// TIA Portal project "Factory_Project_V17" (V17)
// Vorlageprojekt für das Buch mit Zielsystem S7-1200

(* hardware
DEVICE "S7-1200-Station_1"  S7-1200 Station
   slot 0: "Baugruppenträger_0"  Rack  V1.0
   slot 1: "PLC_1"  CPU 1211C DC/DC/DC  6ES7 211-1AE40-0XB0  V4.1
DEVICE "HMI_1"  KTP700 Basic PN
   slot 0: "HMI_1"  KTP700 Basic PN  6AV2 123-2GB03-0AX0  17.0.0.0
   slot 1: "HMI_RT_1"  KTP700 Basic PN  6AV2 123-2GB03-0AX0  17.0.0.0
   slot 5: "HMI_1.IE_CP_1"  PROFINET Interface  17.0.0.0
      slot 1: "PROFINET Interface_1"  PROFINET Interface
         slot 1: "Port_1"  Port
*)

// ===== PLC "PLC_1"  CPU 1211C DC/DC/DC =====

VAR_GLOBAL   // PLC tag table "Standard-Variablentabelle"
   "Tag_4" AT %M0.0 : Bool;
   "Tag_5" AT %M0.1 : Bool;
   "Tag_1" AT %M0.3 : Bool;
   "Tag_2" AT %M0.4 : Bool;
   "Tag_3" AT %M100.0 : Bool;
   "Tag_6" AT %M100.1 : Bool;
   "Tag_7" AT %M100.2 : Bool;
   "Tag_8" AT %M100.3 : Bool;
   "Tag_9" AT %M100.4 : Bool;
   "Tag_10" AT %M100.5 : Bool;
   "Tag_11" AT %M100.6 : Bool;
   "Tag_12" AT %M100.7 : Bool;
END_VAR

VAR_GLOBAL   // PLC tag table "Inputs_Tags"
   "start" AT %I0.0 : Bool;
   "stop" AT %I0.1 : Bool;
   "reset" AT %I0.2 : Bool;
   "emergency" AT %I0.3 : Bool;
   "Z1_Presence_sensor" AT %I0.4 : Bool;
   "at_scale_sensor" AT %I0.5 : Bool;
   "Z1_vision_sensor" AT %I0.6 : Bool;
   "machine A entry sensor" AT %I0.7 : Bool;
   "machine B entry sensor" AT %I1.0 : Bool;
   "machine A exit sensor" AT %I1.1 : Bool;
   "machine B exit sensor" AT %I1.2 : Bool;
   "machine A has error" AT %I1.3 : Bool;
   "machine A is busy" AT %I1.4 : Bool;
   "machine A opened" AT %I1.5 : Bool;
   "machine B has error" AT %I1.6 : Bool;
   "machine B is busy" AT %I1.7 : Bool;
   "machine B opened" AT %I2.0 : Bool;
   "up elevator A right limit" AT %I2.1 : Bool;
   "up elevator A left limit" AT %I2.2 : Bool;
   "down elevator A right limit" AT %I2.3 : Bool;
   "down elevator A left limit" AT %I2.4 : Bool;
   "up elevator B right limit" AT %I2.5 : Bool;
   "up elevator B left limit" AT %I2.6 : Bool;
   "down elevator B right limit" AT %I2.7 : Bool;
   "down elevator B left limit" AT %I3.0 : Bool;
   "product A at assemply" AT %I3.3 : Bool;
   "product B at assemply" AT %I3.4 : Bool;
   "product left assemply" AT %I3.5 : Bool;
   "positioner A limit" AT %I3.6 : Bool;
   "positioner A clamped" AT %I3.7 : Bool;
   "positioner B limit" AT %I4.0 : Bool;
   "Positioner B clamped" AT %I4.1 : Bool;
   "assempler moving x" AT %I4.2 : Bool;
   "assempler  moving z" AT %I4.3 : Bool;
   "assempler rotating" AT %I4.4 : Bool;
   "assempler item detected" AT %I4.5 : Bool;
   "assempler gripper rotating" AT %I4.6 : Bool;
   "palletizer elevator back limit" AT %I4.7 : Bool;
   "palletizer elevator front limit" AT %I5.0 : Bool;
   "palletizer clamped" AT %I5.1 : Bool;
   "palletizer elevator moving" AT %I5.2 : Bool;
   "palletizer plate limit" AT %I5.3 : Bool;
   "palletizer pusher limit" AT %I5.4 : Bool;
   "stacker crane moving x" AT %I5.5 : Bool;
   "stacker crane moving z" AT %I5.6 : Bool;
   "stacker crane left limit" AT %I5.7 : Bool;
   "stacker crane right limit" AT %I6.0 : Bool;
   "stacker crane middle limit" AT %I6.1 : Bool;
   "scale value" AT %ID32 : Real;
   "UP ELEVATOR A POSITION" AT %ID36 : Real;
   "DOWN ELEVATOR A POSITION" AT %ID40 : Real;
   "assempler position x" AT %ID44 : Real;
   "assempler position z" AT %ID48 : Real;
   "bridge A1 sensor" AT %I6.2 : Bool;
   "bridge A2 sensor" AT %I6.3 : Bool;
   "bridge B1 sensor" AT %I6.4 : Bool;
   "bridge B2 sensor" AT %I6.5 : Bool;
   "UP ELEVATOR B POSITION" AT %ID52 : Real;
   "DOWN ELEVATOR B POSITION" AT %ID56 : Real;
   "PALLETIZER ENTRY" AT %I6.6 : Bool;
   "LOADING CONV ENTRY SENSOR" AT %I6.7 : Bool;
   "LOADING CONV EXIT SENSOR" AT %I7.0 : Bool;
END_VAR

VAR_GLOBAL   // PLC tag table "Outputs_tags"
   "start light" AT %Q0.0 : Bool;
   "stop light" AT %Q0.1 : Bool;
   "reset light" AT %Q0.2 : Bool;
   "error light 1" AT %Q0.3 : Bool;
   "error light 2" AT %Q0.4 : Bool;
   "warning light 1" AT %Q0.5 : Bool;
   "warning light 2" AT %Q0.6 : Bool;
   "feed conv" AT %Q0.7 : Bool;
   "feed emittor" AT %Q1.0 : Bool;
   "scale conv" AT %Q1.1 : Bool;
   "sorter wheels" AT %Q1.2 : Bool;
   "sorter right" AT %Q1.3 : Bool;
   "sorter left" AT %Q1.4 : Bool;
   "Z1L1" AT %Q1.5 : Bool;
   "Z1L2" AT %Q1.6 : Bool;
   "Z1L3" AT %Q1.7 : Bool;
   "Z1L4" AT %Q2.0 : Bool;
   "Z1L5" AT %Q2.1 : Bool;
   "Z1L6" AT %Q2.2 : Bool;
   "Z1L7" AT %Q2.3 : Bool;
   "Z1L8" AT %Q2.4 : Bool;
   "Z1R1" AT %Q2.5 : Bool;
   "Z1R2" AT %Q2.6 : Bool;
   "Z1R3" AT %Q2.7 : Bool;
   "Z1R4" AT %Q3.0 : Bool;
   "Z1R5" AT %Q3.1 : Bool;
   "Z1R6" AT %Q3.2 : Bool;
   "Z3A1" AT %Q3.3 : Bool;
   "Z3A2" AT %Q3.4 : Bool;
   "Z3A3" AT %Q3.5 : Bool;
   "Z3A4" AT %Q3.6 : Bool;
   "Z3A5" AT %Q3.7 : Bool;
   "Z3A6" AT %Q4.0 : Bool;
   "Z3B1" AT %Q4.1 : Bool;
   "Z3B2" AT %Q4.2 : Bool;
   "Z3B3" AT %Q4.3 : Bool;
   "Z3B4" AT %Q4.4 : Bool;
   "Z3B5" AT %Q4.5 : Bool;
   "Z3B6" AT %Q4.6 : Bool;
   "Z3B7" AT %Q4.7 : Bool;
   "Z4_1" AT %Q5.2 : Bool;
   "Z4_2" AT %Q5.3 : Bool;
   "Z4_3" AT %Q5.4 : Bool;
   "Z4_4" AT %Q5.5 : Bool;
   "Z4 entry roller" AT %Q5.7 : Bool;
   "Z4 exit roller" AT %Q6.0 : Bool;
   "loading entry conv" AT %Q6.1 : Bool;
   "loading exit conv" AT %Q6.2 : Bool;
   "exit conv 1" AT %Q6.3 : Bool;
   "exit conv 2" AT %Q6.4 : Bool;
   "exit conv 3" AT %Q6.5 : Bool;
   "machine A start" AT %Q6.6 : Bool;
   "machine A stop" AT %Q6.7 : Bool;
   "machine A reset" AT %Q7.0 : Bool;
   "machine A lids" AT %Q7.1 : Bool;
   "machine B start" AT %Q7.2 : Bool;
   "Z4_5" AT %Q5.6 : Bool;
   "machine B stop" AT %Q7.3 : Bool;
   "machine B reset" AT %Q7.4 : Bool;
   "machine B lids" AT %Q7.5 : Bool;
   "up elevator A +" AT %Q7.6 : Bool;
   "up elevator A -" AT %Q7.7 : Bool;
   "up elevator A stop blade" AT %Q8.0 : Bool;
   "up elevator B +" AT %Q8.1 : Bool;
   "up elevator B -" AT %Q8.2 : Bool;
   "up elevator B stop blade" AT %Q8.3 : Bool;
   "down elevator A +" AT %Q8.4 : Bool;
   "down elevator A -" AT %Q8.5 : Bool;
   "down elevator A stop blade" AT %Q8.6 : Bool;
   "down elevator B+" AT %Q8.7 : Bool;
   "down elevator B -" AT %Q9.0 : Bool;
   "down elevator B stop blade" AT %Q9.1 : Bool;
   "positioner A raise" AT %Q9.2 : Bool;
   "positioner A clamp" AT %Q9.3 : Bool;
   "positioner B raise" AT %Q9.4 : Bool;
   "positioner B clamp" AT %Q9.5 : Bool;
   "assempler grap" AT %Q9.6 : Bool;
   "assempler rotate cw" AT %Q9.7 : Bool;
   "assempler rotate ccw" AT %Q10.1 : Bool;
   "assempler gripper ccw" AT %Q10.2 : Bool;
   "palletizer turn" AT %Q10.3 : Bool;
   "palletizer push" AT %Q10.4 : Bool;
   "palletizer clamp" AT %Q10.5 : Bool;
   "palletizer open plate" AT %Q10.6 : Bool;
   "palletizer belt +" AT %Q10.7 : Bool;
   "palletizer belt -" AT %Q11.0 : Bool;
   "palletizer chain +" AT %Q11.1 : Bool;
   "palletizer chain -" AT %Q11.2 : Bool;
   "palletizer elevator +" AT %Q11.3 : Bool;
   "palletizer elevator -" AT %Q11.4 : Bool;
   "palletizer elevator move to limit" AT %Q11.5 : Bool;
   "stacker crane lift" AT %Q11.6 : Bool;
   "stacker crane left" AT %Q11.7 : Bool;
   "stacker crane right" AT %Q12.0 : Bool;
   "state" AT %QD32 : DInt;
   "up elevator A set point" AT %QD36 : Real;
   "up elevator B set point" AT %QD40 : Real;
   "down elevator A set point" AT %QD44 : Real;
   "down elevator B set point" AT %QD48 : Real;
   "assempler x set point" AT %QD52 : Real;
   "assempler z set point" AT %QD56 : Real;
   "stacker crane target position" AT %QD60 : DInt;
   "bridge A1 stop blade" AT %Q12.1 : Bool;
   "bridge A2 stop blade" AT %Q12.2 : Bool;
   "bridge B1 stop blade" AT %Q12.3 : Bool;
   "bridge B2 stop blade" AT %Q12.4 : Bool;
   "Z3-A1 bridge conv" AT %Q12.5 : Bool;
   "Z3-A2 bridge conv" AT %Q12.6 : Bool;
   "Z3-A3 bridge conv" AT %Q12.7 : Bool;
   "Z3-B1 bridge conv" AT %Q13.0 : Bool;
   "Z3-B2 bridge conv" AT %Q13.1 : Bool;
   "Z3-B3 bridge conv" AT %Q13.2 : Bool;
   "PALLETIZER EMITTER" AT %Q10.0 : Bool;
END_VAR

VAR_GLOBAL   // PLC tag table "alarm_tags"
   "Alarm_trigger" AT %MW100 : Word;
END_VAR

TYPE "RackSlot"
   STRUCT
      occupied : Bool;
      side : Int;
      space : Int;
   END_STRUCT;
END_TYPE

DATA_BLOCK "DB_RackMemory"   // DB8
{ S7_Optimized_Access := 'TRUE' }
VERSION : 0.1
   VAR
      Rack : Array[1..108] of "RackSlot";
      SpacesOccupied : Int;
      "FREE SPACES" : Int;
      "QUANTITY TO RETRIEVE" : Int;
      "REQUIRED QUANTITY" : Int;
      RETRIEVE : Bool;
      In_Production : Int;
      "TOTAL ORDERS" : Int;
      "TOTAL DLIEVERED" : Int;
      ReckMemoryReset : Bool;
      InProductionReset : Bool;
   END_VAR
BEGIN
END_DATA_BLOCK

DATA_BLOCK "DB_HMI"   // DB10
{ S7_Optimized_Access := 'TRUE' }
VERSION : 0.1
   VAR
      "Z1 STATUS" : Int;
      "Z2 STATUS" : Int;
      "Z3 BUFFER A STATUS" : Int;
      "Z3 BUFFER B STATUS" : Int;
      "Z3 ASSEMPLER STATUS" : Int;
      "Z4 UPPER STATUS" : Int;
      "Z4 LOWER STATUS" : Int;
      "Z5 STATUS" : Int;
      "FACTORY STATUS" : Int;
      "ASSEMPLER X" : Real;
      "ASSEMPLER Z" : Real;
      "ASSEMPLER GRAB" : Bool;
      "ASSEMPLER ROT CW" : Bool;
      "ASSEMPLER ROT CCW" : Bool;
      "CRANE TARGET" : Int;
      "CRANE SIDE" : Int;
      "CRANE LEFT" : Bool;
      "CRANE LIFT" : Bool;
      "CRANE RIGHT" : Bool;
      "CREATE ORDER" : Bool;
      "CANCEL ORDER" : Bool;
      "MAINTENANCE MODE" : Bool;
      ACK : Bool;
   END_VAR
BEGIN
END_DATA_BLOCK

DATA_BLOCK "FACTORY STATUS MANAGMENT_DB"   // DB11
{ S7_Optimized_Access := 'TRUE' }
VERSION : 0.1
// stored: InstanceOfName FACTORY STATUS MANAGMENT
"FACTORY STATUS MANAGMENT"
BEGIN
END_DATA_BLOCK

// folder: System blocks/Program resources

DATA_BLOCK "z1_timer_ton"   // DB3
{ S7_Optimized_Access := 'TRUE' }
AUTHOR : Simatic
FAMILY : IEC
NAME : IEC_TMR
VERSION : 1.0
// stored: InstanceOfName IEC_TIMER
"IEC_TIMER"
BEGIN
END_DATA_BLOCK

// folder: ZONE-5-BLOCKS

DATA_BLOCK "ZONE-5-FB_DB"   // DB9
{ S7_Optimized_Access := 'TRUE' }
VERSION : 0.1
// stored: InstanceOfName ZONE-5-FB
"ZONE-5-FB"
BEGIN
END_DATA_BLOCK

// folder: ZONE_1_BLOCKS

DATA_BLOCK "Zone_1_FB_DB"   // DB2
{ S7_Optimized_Access := 'TRUE' }
VERSION : 0.1
// stored: InstanceOfName Zone_1_FB
"Zone_1_FB"
BEGIN
END_DATA_BLOCK

// folder: ZONE_4_BLOCKS

DATA_BLOCK "ZONE 4 FB_DB"   // DB7
{ S7_Optimized_Access := 'TRUE' }
VERSION : 0.1
// stored: InstanceOfName ZONE 4 FB
"ZONE 4 FB"
BEGIN
END_DATA_BLOCK

// folder: Zone _2_Blocks

DATA_BLOCK "Zone_2_FB_DB"   // DB4
{ S7_Optimized_Access := 'TRUE' }
VERSION : 0.1
// stored: InstanceOfName Zone_2_FB
"Zone_2_FB"
BEGIN
END_DATA_BLOCK

// folder: Zone_3_blocks

DATA_BLOCK "Zone_3_FB_DB"   // DB5
{ S7_Optimized_Access := 'TRUE' }
VERSION : 0.1
// stored: InstanceOfName Zone_3_FB
"Zone_3_FB"
BEGIN
END_DATA_BLOCK

// folder: Zone_3_blocks/BUFFER SUB BLOCKS

DATA_BLOCK "ZONE-3 BUFFER_A_DB"   // DB6
{ S7_Optimized_Access := 'TRUE' }
VERSION : 0.1
// stored: InstanceOfName ZONE-3 BUFFER
"ZONE-3 BUFFER"
BEGIN
END_DATA_BLOCK

// folder: (top level)

FUNCTION_BLOCK "FACTORY STATUS MANAGMENT"   // FB22, SCL
{ S7_Optimized_Access := 'TRUE' }
VERSION : 0.1
   VAR_INPUT
      START : Bool;
      STOP : Bool;
      RESET : Bool;
      "Z1 STATUS" : Int;
      "Z2 STATUS" : Int;
      "Z3 BUFFER A STATUS" : Int;
      "Z3 BUFFER B STATUS" : Int;
      "Z3 ASSEMPLER STATUS" : Int;
      "Z4 STATUS UPPER" : Int;
      "Z4 LOWER STATUS" : Int;
      "Z5 STATUS" : Int;
   END_VAR
   VAR_OUTPUT
      "FACTORY STATUS" : Int;
   END_VAR
BEGIN
   IF #"Z1 STATUS" = 90
       OR #"Z2 STATUS" = 90
       OR #"Z3 BUFFER A STATUS" = 90
       OR #"Z3 BUFFER B STATUS" = 90
       OR #"Z3 ASSEMPLER STATUS" = 90
       OR #"Z4 STATUS UPPER" = 90
       OR #"Z4 LOWER STATUS" = 90
       OR #"Z5 STATUS" = 90
   THEN
       #"FACTORY STATUS" := 90;
   END_IF;

   IF #"FACTORY STATUS" = 90 THEN
       IF #RESET THEN
           #"FACTORY STATUS" := 0;
       END_IF;
   END_IF;

   IF #START AND  #"FACTORY STATUS" <> 90 THEN
       #"FACTORY STATUS" := 10;
   END_IF;

   IF #STOP AND #"FACTORY STATUS" <> 90 THEN
       #"FACTORY STATUS" := 0;
   END_IF;
END_FUNCTION_BLOCK

FUNCTION "MHJ-PLC-Lab-Function-S71200" : Void   // FC9000, SCL
{ S7_Optimized_Access := 'TRUE' }
VERSION : 0.1
   VAR_TEMP
      rdTimeReturn : Int;
      outputTime : DTL;
      SyncVal : Byte;
      forVal : Int;
      forVal_2 : Int;
      Value : Byte;
   END_VAR
   VAR CONSTANT
      CompVal : Byte := 16#34;
      Value_01 : Byte := 16#11;
      Value_01_DW : DWord := 16#A165_D992;
      Value_02_DW : DWord := 16#58BE_4401;
   END_VAR
BEGIN

   #Value:=PEEK(area := 16#82,
        dbNumber := 0,
        byteOffset := 511);
   #Value := #Value + 1;

   POKE(area := 16#82,
        dbNumber := 0,
        byteOffset := 511,
        value := #Value);

   POKE(area:=16#81,
        dbNumber:=0,
        byteOffset:=1016,
        value:=#Value_01_DW);
   POKE(area := 16#81,
        dbNumber := 0,
        byteOffset := 1020,
        value := #Value_02_DW);

   POKE(area := 16#81,
        dbNumber := 0,
        byteOffset := 511,
        value := B#16#00);

   FOR #forVal := 0 TO 120 DO
       FOR #forVal_2:=0 TO 10 DO
           #rdTimeReturn:=RD_SYS_T(#outputTime);
           #rdTimeReturn := WR_SYS_T(#outputTime);
           #rdTimeReturn := RD_SYS_T(#outputTime);
           #rdTimeReturn := WR_SYS_T(#outputTime);
       END_FOR;
       #SyncVal:= PEEK(area := 16#81,
                      dbNumber := 0,
                      byteOffset := 511);
       IF #SyncVal = #CompVal THEN
          GOTO M_1;
       END_IF;
   END_FOR;
   RETURN;

   M_1:
   POKE(area := 16#81,
        dbNumber := 0,
        byteOffset := 511,
        value := B#16#0);
END_FUNCTION

ORGANIZATION_BLOCK "Main"   // OB1, LAD, ProgramCycle
TITLE = "Main Program Sweep (Cycle)"
{ S7_Optimized_Access := 'TRUE' }
VERSION : 0.1
   VAR_INPUT
      Initial_Call : Bool;   // Initial call of this OB
      Remanence : Bool;   // =True, if remanent data are available
   END_VAR
BEGIN

REGION Network 1: Konnektierungsbaustein für PLC-Lab
   // Im Netzwerk 1 wird der Konnektierungsbaustein für PLC-Lab aufgerufen.
   // Dieser Aufruf darf nicht entfernt werden!
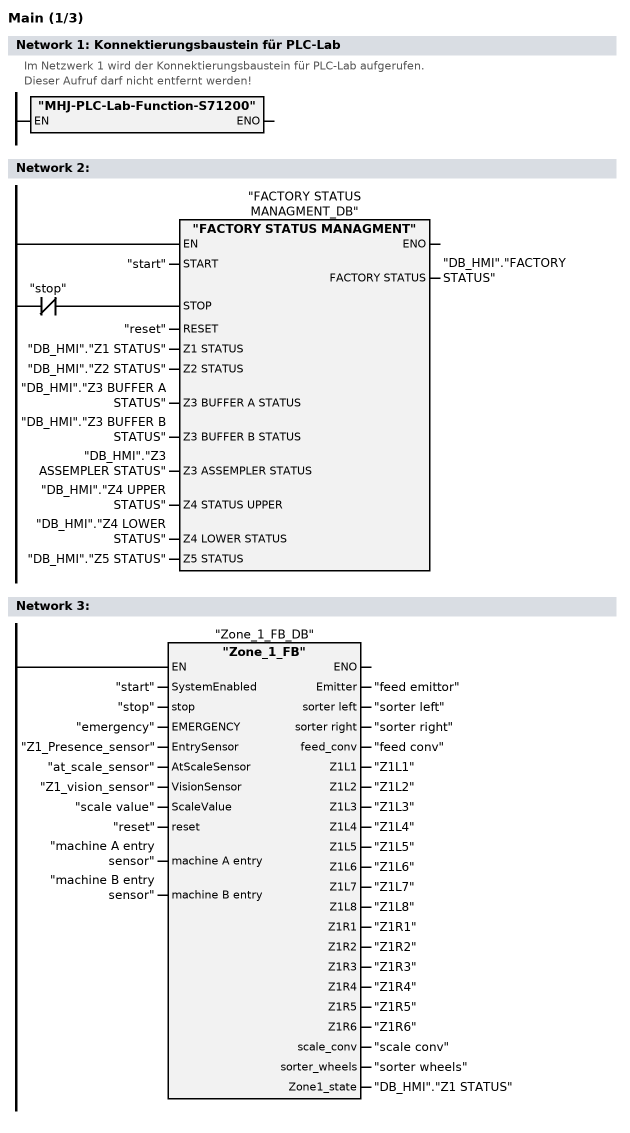
   RUNG wire#powerrail
      "MHJ-PLC-Lab-Function-S71200"()
   END_RUNG
   // the same network as SCL:
   "MHJ-PLC-Lab-Function-S71200"();
END_REGION

REGION Network 2
   RUNG wire#powerrail
      "FACTORY STATUS MANAGMENT_DB"(STOP := wire#w1, START := "start", RESET := "reset", "Z1 STATUS" := "DB_HMI"."Z1 STATUS", "Z2 STATUS" := "DB_HMI"."Z2 STATUS", "Z3 BUFFER A STATUS" := "DB_HMI"."Z3 BUFFER A STATUS", "Z3 BUFFER B STATUS" := "DB_HMI"."Z3 BUFFER B STATUS", "Z3 ASSEMPLER STATUS" := "DB_HMI"."Z3 ASSEMPLER STATUS", "Z4 STATUS UPPER" := "DB_HMI"."Z4 UPPER STATUS", "Z4 LOWER STATUS" := "DB_HMI"."Z4 LOWER STATUS", "Z5 STATUS" := "DB_HMI"."Z5 STATUS", "FACTORY STATUS" => "DB_HMI"."FACTORY STATUS")
   END_RUNG
   RUNG wire#powerrail
      I_Contact( "stop" )
   END_RUNG wire#w1
   // the same network as SCL:
   "FACTORY STATUS MANAGMENT_DB"(START := "start",   // "FACTORY STATUS MANAGMENT"
                           STOP := NOT "stop",
                           RESET := "reset",
                           "Z1 STATUS" := "DB_HMI"."Z1 STATUS",
                           "Z2 STATUS" := "DB_HMI"."Z2 STATUS",
                           "Z3 BUFFER A STATUS" := "DB_HMI"."Z3 BUFFER A STATUS",
                           "Z3 BUFFER B STATUS" := "DB_HMI"."Z3 BUFFER B STATUS",
                           "Z3 ASSEMPLER STATUS" := "DB_HMI"."Z3 ASSEMPLER STATUS",
                           "Z4 STATUS UPPER" := "DB_HMI"."Z4 UPPER STATUS",
                           "Z4 LOWER STATUS" := "DB_HMI"."Z4 LOWER STATUS",
                           "Z5 STATUS" := "DB_HMI"."Z5 STATUS",
                           "FACTORY STATUS" => "DB_HMI"."FACTORY STATUS");
END_REGION

REGION Network 3
   RUNG wire#powerrail
      "Zone_1_FB_DB"(SystemEnabled := "start", stop := "stop", EMERGENCY := "emergency", EntrySensor := "Z1_Presence_sensor", AtScaleSensor := "at_scale_sensor", VisionSensor := "Z1_vision_sensor", ScaleValue := "scale value", reset := "reset", "machine A entry" := "machine A entry sensor", "machine B entry" := "machine B entry sensor", Emitter => "feed emittor", "sorter left" => "sorter left", "sorter right" => "sorter right", feed_conv => "feed conv", Z1L1 => "Z1L1", Z1L2 => "Z1L2", Z1L3 => "Z1L3", Z1L4 => "Z1L4", Z1L5 => "Z1L5", Z1L6 => "Z1L6", Z1L7 => "Z1L7", Z1L8 => "Z1L8", Z1R1 => "Z1R1", Z1R2 => "Z1R2", Z1R3 => "Z1R3", Z1R4 => "Z1R4", Z1R5 => "Z1R5", Z1R6 => "Z1R6", scale_conv => "scale conv", sorter_wheels => "sorter wheels", Zone1_state => "DB_HMI"."Z1 STATUS")
   END_RUNG
   // the same network as SCL:
   "Zone_1_FB_DB"(SystemEnabled := "start",   // "Zone_1_FB"
                  stop := "stop",
                  EMERGENCY := "emergency",
                  EntrySensor := "Z1_Presence_sensor",
                  AtScaleSensor := "at_scale_sensor",
                  VisionSensor := "Z1_vision_sensor",
                  ScaleValue := "scale value",
                  reset := "reset",
                  "machine A entry" := "machine A entry sensor",
                  "machine B entry" := "machine B entry sensor",
                  Emitter => "feed emittor",
                  "sorter left" => "sorter left",
                  "sorter right" => "sorter right",
                  feed_conv => "feed conv",
                  Z1L1 => "Z1L1",
                  Z1L2 => "Z1L2",
                  Z1L3 => "Z1L3",
                  Z1L4 => "Z1L4",
                  Z1L5 => "Z1L5",
                  Z1L6 => "Z1L6",
                  Z1L7 => "Z1L7",
                  Z1L8 => "Z1L8",
                  Z1R1 => "Z1R1",
                  Z1R2 => "Z1R2",
                  Z1R3 => "Z1R3",
                  Z1R4 => "Z1R4",
                  Z1R5 => "Z1R5",
                  Z1R6 => "Z1R6",
                  scale_conv => "scale conv",
                  sorter_wheels => "sorter wheels",
                  Zone1_state => "DB_HMI"."Z1 STATUS");
END_REGION

REGION Network 4
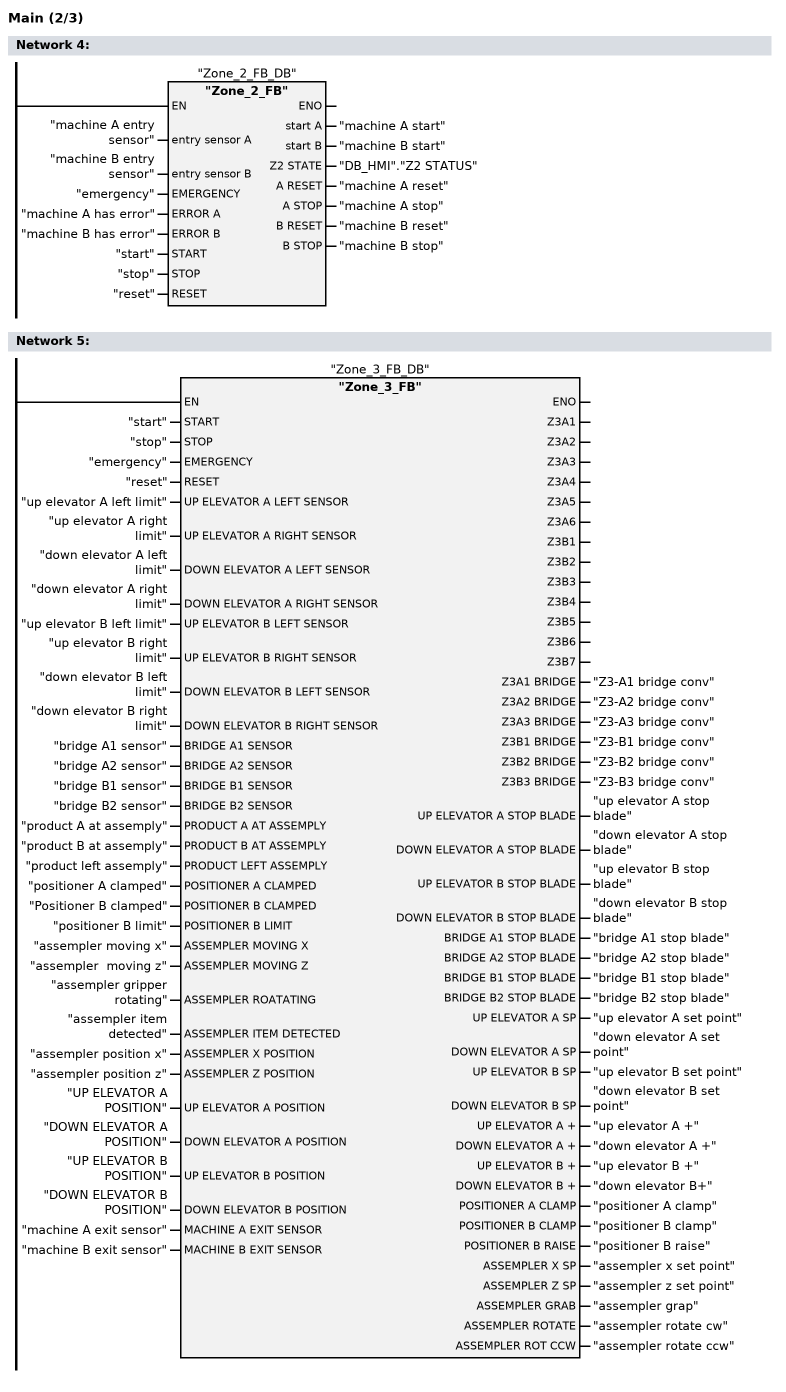
   RUNG wire#powerrail
      "Zone_2_FB_DB"("entry sensor A" := "machine A entry sensor", "entry sensor B" := "machine B entry sensor", EMERGENCY := "emergency", "ERROR A" := "machine A has error", "ERROR B" := "machine B has error", START := "start", STOP := "stop", RESET := "reset", "start A" => "machine A start", "start B" => "machine B start", "Z2 STATE" => "DB_HMI"."Z2 STATUS", "A RESET" => "machine A reset", "A STOP" => "machine A stop", "B RESET" => "machine B reset", "B STOP" => "machine B stop")
   END_RUNG
   // the same network as SCL:
   "Zone_2_FB_DB"("entry sensor A" := "machine A entry sensor",   // "Zone_2_FB"
                  "entry sensor B" := "machine B entry sensor",
                  EMERGENCY := "emergency",
                  "ERROR A" := "machine A has error",
                  "ERROR B" := "machine B has error",
                  START := "start",
                  STOP := "stop",
                  RESET := "reset",
                  "start A" => "machine A start",
                  "start B" => "machine B start",
                  "Z2 STATE" => "DB_HMI"."Z2 STATUS",
                  "A RESET" => "machine A reset",
                  "A STOP" => "machine A stop",
                  "B RESET" => "machine B reset",
                  "B STOP" => "machine B stop");
END_REGION

REGION Network 5
   RUNG wire#powerrail
      "Zone_3_FB_DB"(START := "start", STOP := "stop", EMERGENCY := "emergency", RESET := "reset", "UP ELEVATOR A LEFT SENSOR" := "up elevator A left limit", "UP ELEVATOR A RIGHT SENSOR" := "up elevator A right limit", "DOWN ELEVATOR A LEFT SENSOR" := "down elevator A left limit", "DOWN ELEVATOR A RIGHT SENSOR" := "down elevator A right limit", "UP ELEVATOR B LEFT SENSOR" := "up elevator B left limit", "UP ELEVATOR B RIGHT SENSOR" := "up elevator B right limit", "DOWN ELEVATOR B LEFT SENSOR" := "down elevator B left limit", "DOWN ELEVATOR B RIGHT SENSOR" := "down elevator B right limit", "BRIDGE A1 SENSOR" := "bridge A1 sensor", "BRIDGE A2 SENSOR" := "bridge A2 sensor", "BRIDGE B1 SENSOR" := "bridge B1 sensor", "BRIDGE B2 SENSOR" := "bridge B2 sensor", "PRODUCT A AT ASSEMPLY" := "product A at assemply", "PRODUCT B AT ASSEMPLY" := "product B at assemply", "PRODUCT LEFT ASSEMPLY" := "product left assemply", "POSITIONER A CLAMPED" := "positioner A clamped", "POSITIONER B CLAMPED" := "Positioner B clamped", "POSITIONER B LIMIT" := "positioner B limit", "ASSEMPLER MOVING X" := "assempler moving x", "ASSEMPLER MOVING Z" := "assempler  moving z", "ASSEMPLER ROATATING" := "assempler gripper rotating", "ASSEMPLER ITEM DETECTED" := "assempler item detected", "ASSEMPLER X POSITION" := "assempler position x", "ASSEMPLER Z POSITION" := "assempler position z", "UP ELEVATOR A POSITION" := "UP ELEVATOR A POSITION", "DOWN ELEVATOR A POSITION" := "DOWN ELEVATOR A POSITION", "UP ELEVATOR B POSITION" := "UP ELEVATOR B POSITION", "DOWN ELEVATOR B POSITION" := "DOWN ELEVATOR B POSITION", "MACHINE A EXIT SENSOR" := "machine A exit sensor", "MACHINE B EXIT SENSOR" := "machine B exit sensor", Z3A1 =>, Z3A2 =>, Z3A3 =>, Z3A4 =>, Z3A5 =>, Z3A6 =>, Z3B1 =>, Z3B2 =>, Z3B3 =>, Z3B4 =>, Z3B5 =>, Z3B6 =>, Z3B7 =>, "Z3A1 BRIDGE" => "Z3-A1 bridge conv", "Z3A2 BRIDGE" => "Z3-A2 bridge conv", "Z3A3 BRIDGE" => "Z3-A3 bridge conv", "Z3B1 BRIDGE" => "Z3-B1 bridge conv", "Z3B2 BRIDGE" => "Z3-B2 bridge conv", "Z3B3 BRIDGE" => "Z3-B3 bridge conv", "UP ELEVATOR A STOP BLADE" => "up elevator A stop blade", "DOWN ELEVATOR A STOP BLADE" => "down elevator A stop blade", "UP ELEVATOR B STOP BLADE" => "up elevator B stop blade", "DOWN ELEVATOR B STOP BLADE" => "down elevator B stop blade", "BRIDGE A1 STOP BLADE" => "bridge A1 stop blade", "BRIDGE A2 STOP BLADE" => "bridge A2 stop blade", "BRIDGE B1 STOP BLADE" => "bridge B1 stop blade", "BRIDGE B2 STOP BLADE" => "bridge B2 stop blade", "UP ELEVATOR A SP" => "up elevator A set point", "DOWN ELEVATOR A SP" => "down elevator A set point", "UP ELEVATOR B SP" => "up elevator B set point", "DOWN ELEVATOR B SP" => "down elevator B set point", "UP ELEVATOR A +" => "up elevator A +", "DOWN ELEVATOR A +" => "down elevator A +", "UP ELEVATOR B +" => "up elevator B +", "DOWN ELEVATOR B +" => "down elevator B+", "POSITIONER A CLAMP" => "positioner A clamp", "POSITIONER B CLAMP" => "positioner B clamp", "POSITIONER B RAISE" => "positioner B raise", "ASSEMPLER X SP" => "assempler x set point", "ASSEMPLER Z SP" => "assempler z set point", "ASSEMPLER GRAB" => "assempler grap", "ASSEMPLER ROTATE" => "assempler rotate cw", "ASSEMPLER ROT CCW" => "assempler rotate ccw")
   END_RUNG
   // the same network as SCL:
   "Zone_3_FB_DB"(START := "start",   // "Zone_3_FB"
                  STOP := "stop",
                  EMERGENCY := "emergency",
                  RESET := "reset",
                  "UP ELEVATOR A LEFT SENSOR" := "up elevator A left limit",
                  "UP ELEVATOR A RIGHT SENSOR" := "up elevator A right limit",
                  "DOWN ELEVATOR A LEFT SENSOR" := "down elevator A left limit",
                  "DOWN ELEVATOR A RIGHT SENSOR" := "down elevator A right limit",
                  "UP ELEVATOR B LEFT SENSOR" := "up elevator B left limit",
                  "UP ELEVATOR B RIGHT SENSOR" := "up elevator B right limit",
                  "DOWN ELEVATOR B LEFT SENSOR" := "down elevator B left limit",
                  "DOWN ELEVATOR B RIGHT SENSOR" := "down elevator B right limit",
                  "BRIDGE A1 SENSOR" := "bridge A1 sensor",
                  "BRIDGE A2 SENSOR" := "bridge A2 sensor",
                  "BRIDGE B1 SENSOR" := "bridge B1 sensor",
                  "BRIDGE B2 SENSOR" := "bridge B2 sensor",
                  "PRODUCT A AT ASSEMPLY" := "product A at assemply",
                  "PRODUCT B AT ASSEMPLY" := "product B at assemply",
                  "PRODUCT LEFT ASSEMPLY" := "product left assemply",
                  "POSITIONER A CLAMPED" := "positioner A clamped",
                  "POSITIONER B CLAMPED" := "Positioner B clamped",
                  "POSITIONER B LIMIT" := "positioner B limit",
                  "ASSEMPLER MOVING X" := "assempler moving x",
                  "ASSEMPLER MOVING Z" := "assempler  moving z",
                  "ASSEMPLER ROATATING" := "assempler gripper rotating",
                  "ASSEMPLER ITEM DETECTED" := "assempler item detected",
                  "ASSEMPLER X POSITION" := "assempler position x",
                  "ASSEMPLER Z POSITION" := "assempler position z",
                  "UP ELEVATOR A POSITION" := "UP ELEVATOR A POSITION",
                  "DOWN ELEVATOR A POSITION" := "DOWN ELEVATOR A POSITION",
                  "UP ELEVATOR B POSITION" := "UP ELEVATOR B POSITION",
                  "DOWN ELEVATOR B POSITION" := "DOWN ELEVATOR B POSITION",
                  "MACHINE A EXIT SENSOR" := "machine A exit sensor",
                  "MACHINE B EXIT SENSOR" := "machine B exit sensor",
                  "Z3A1 BRIDGE" => "Z3-A1 bridge conv",
                  "Z3A2 BRIDGE" => "Z3-A2 bridge conv",
                  "Z3A3 BRIDGE" => "Z3-A3 bridge conv",
                  "Z3B1 BRIDGE" => "Z3-B1 bridge conv",
                  "Z3B2 BRIDGE" => "Z3-B2 bridge conv",
                  "Z3B3 BRIDGE" => "Z3-B3 bridge conv",
                  "UP ELEVATOR A STOP BLADE" => "up elevator A stop blade",
                  "DOWN ELEVATOR A STOP BLADE" => "down elevator A stop blade",
                  "UP ELEVATOR B STOP BLADE" => "up elevator B stop blade",
                  "DOWN ELEVATOR B STOP BLADE" => "down elevator B stop blade",
                  "BRIDGE A1 STOP BLADE" => "bridge A1 stop blade",
                  "BRIDGE A2 STOP BLADE" => "bridge A2 stop blade",
                  "BRIDGE B1 STOP BLADE" => "bridge B1 stop blade",
                  "BRIDGE B2 STOP BLADE" => "bridge B2 stop blade",
                  "UP ELEVATOR A SP" => "up elevator A set point",
                  "DOWN ELEVATOR A SP" => "down elevator A set point",
                  "UP ELEVATOR B SP" => "up elevator B set point",
                  "DOWN ELEVATOR B SP" => "down elevator B set point",
                  "UP ELEVATOR A +" => "up elevator A +",
                  "DOWN ELEVATOR A +" => "down elevator A +",
                  "UP ELEVATOR B +" => "up elevator B +",
                  "DOWN ELEVATOR B +" => "down elevator B+",
                  "POSITIONER A CLAMP" => "positioner A clamp",
                  "POSITIONER B CLAMP" => "positioner B clamp",
                  "POSITIONER B RAISE" => "positioner B raise",
                  "ASSEMPLER X SP" => "assempler x set point",
                  "ASSEMPLER Z SP" => "assempler z set point",
                  "ASSEMPLER GRAB" => "assempler grap",
                  "ASSEMPLER ROTATE" => "assempler rotate cw",
                  "ASSEMPLER ROT CCW" => "assempler rotate ccw");
END_REGION

REGION Network 6
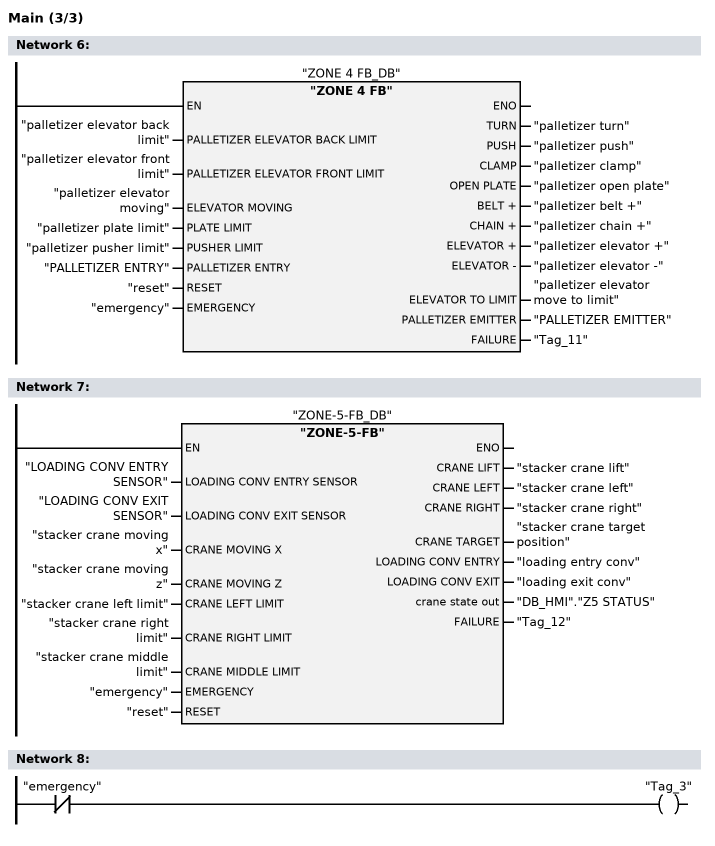
   RUNG wire#powerrail
      "ZONE 4 FB_DB"("PALLETIZER ELEVATOR BACK LIMIT" := "palletizer elevator back limit", "PALLETIZER ELEVATOR FRONT LIMIT" := "palletizer elevator front limit", "ELEVATOR MOVING" := "palletizer elevator moving", "PLATE LIMIT" := "palletizer plate limit", "PUSHER LIMIT" := "palletizer pusher limit", "PALLETIZER ENTRY" := "PALLETIZER ENTRY", RESET := "reset", EMERGENCY := "emergency", TURN => "palletizer turn", PUSH => "palletizer push", CLAMP => "palletizer clamp", "OPEN PLATE" => "palletizer open plate", "BELT +" => "palletizer belt +", "CHAIN +" => "palletizer chain +", "ELEVATOR +" => "palletizer elevator +", "ELEVATOR -" => "palletizer elevator -", "ELEVATOR TO LIMIT" => "palletizer elevator move to limit", "PALLETIZER EMITTER" => "PALLETIZER EMITTER", FAILURE => "Tag_11")
   END_RUNG
   // the same network as SCL:
   "ZONE 4 FB_DB"("PALLETIZER ELEVATOR BACK LIMIT" := "palletizer elevator back limit",   // "ZONE 4 FB"
                  "PALLETIZER ELEVATOR FRONT LIMIT" := "palletizer elevator front limit",
                  "ELEVATOR MOVING" := "palletizer elevator moving",
                  "PLATE LIMIT" := "palletizer plate limit",
                  "PUSHER LIMIT" := "palletizer pusher limit",
                  "PALLETIZER ENTRY" := "PALLETIZER ENTRY",
                  RESET := "reset",
                  EMERGENCY := "emergency",
                  TURN => "palletizer turn",
                  PUSH => "palletizer push",
                  CLAMP => "palletizer clamp",
                  "OPEN PLATE" => "palletizer open plate",
                  "BELT +" => "palletizer belt +",
                  "CHAIN +" => "palletizer chain +",
                  "ELEVATOR +" => "palletizer elevator +",
                  "ELEVATOR -" => "palletizer elevator -",
                  "ELEVATOR TO LIMIT" => "palletizer elevator move to limit",
                  "PALLETIZER EMITTER" => "PALLETIZER EMITTER",
                  FAILURE => "Tag_11");
END_REGION

REGION Network 7
   RUNG wire#powerrail
      "ZONE-5-FB_DB"("LOADING CONV ENTRY SENSOR" := "LOADING CONV ENTRY SENSOR", "LOADING CONV EXIT SENSOR" := "LOADING CONV EXIT SENSOR", "CRANE MOVING X" := "stacker crane moving x", "CRANE MOVING Z" := "stacker crane moving z", "CRANE LEFT LIMIT" := "stacker crane left limit", "CRANE RIGHT LIMIT" := "stacker crane right limit", "CRANE MIDDLE LIMIT" := "stacker crane middle limit", EMERGENCY := "emergency", RESET := "reset", "CRANE LIFT" => "stacker crane lift", "CRANE LEFT" => "stacker crane left", "CRANE RIGHT" => "stacker crane right", "CRANE TARGET" => "stacker crane target position", "LOADING CONV ENTRY" => "loading entry conv", "LOADING CONV EXIT" => "loading exit conv", "crane state out" => "DB_HMI"."Z5 STATUS", FAILURE => "Tag_12")
   END_RUNG
   // the same network as SCL:
   "ZONE-5-FB_DB"("LOADING CONV ENTRY SENSOR" := "LOADING CONV ENTRY SENSOR",   // "ZONE-5-FB"
                  "LOADING CONV EXIT SENSOR" := "LOADING CONV EXIT SENSOR",
                  "CRANE MOVING X" := "stacker crane moving x",
                  "CRANE MOVING Z" := "stacker crane moving z",
                  "CRANE LEFT LIMIT" := "stacker crane left limit",
                  "CRANE RIGHT LIMIT" := "stacker crane right limit",
                  "CRANE MIDDLE LIMIT" := "stacker crane middle limit",
                  EMERGENCY := "emergency",
                  RESET := "reset",
                  "CRANE LIFT" => "stacker crane lift",
                  "CRANE LEFT" => "stacker crane left",
                  "CRANE RIGHT" => "stacker crane right",
                  "CRANE TARGET" => "stacker crane target position",
                  "LOADING CONV ENTRY" => "loading entry conv",
                  "LOADING CONV EXIT" => "loading exit conv",
                  "crane state out" => "DB_HMI"."Z5 STATUS",
                  FAILURE => "Tag_12");
END_REGION

REGION Network 8
   RUNG wire#powerrail
      I_Contact( "emergency" )
      Coil( "Tag_3" )
   END_RUNG
   // the same network as SCL:
   "Tag_3" := NOT "emergency";
END_REGION
END_ORGANIZATION_BLOCK

ORGANIZATION_BLOCK "Startup"   // OB100, SCL, Startup
TITLE = "Complete Restart"
{ S7_Optimized_Access := 'TRUE' }
VERSION : 0.1
   VAR_INPUT
      LostRetentive : Bool;   // True if retentive data are lost
      LostRTC : Bool;   // True if date and time are lost
   END_VAR
   VAR_TEMP
      i : Int;
   END_VAR
BEGIN
   FOR #i := 1 TO 108 DO

       "DB_RackMemory".Rack[#i].occupied := FALSE;

       IF #i <= 54 THEN
           "DB_RackMemory".Rack[#i].side := 1;
           "DB_RackMemory".Rack[#i].space := #i;
       ELSE
           "DB_RackMemory".Rack[#i].side := 2;
           "DB_RackMemory".Rack[#i].space := #i - 54;
       END_IF;

   END_FOR;
END_ORGANIZATION_BLOCK

// folder: ZONE-5-BLOCKS

FUNCTION_BLOCK "ZONE-5-FB"   // FB19, LAD
{ S7_Optimized_Access := 'TRUE' }
VERSION : 0.1
   VAR_INPUT
      "LOADING CONV ENTRY SENSOR" : Bool;
      "LOADING CONV EXIT SENSOR" : Bool;
      "CRANE MOVING X" : Bool;
      "CRANE MOVING Z" : Bool;
      "CRANE LEFT LIMIT" : Bool;
      "CRANE RIGHT LIMIT" : Bool;
      "CRANE MIDDLE LIMIT" : Bool;
      EMERGENCY : Bool;
      RESET : Bool;
   END_VAR
   VAR_OUTPUT
      "CRANE LIFT" : Bool;
      "CRANE LEFT" : Bool;
      "CRANE RIGHT" : Bool;
      "CRANE TARGET" : DInt;
      "LOADING CONV ENTRY" : Bool;
      "LOADING CONV EXIT" : Bool;
      "crane state out" : Int;
      FAILURE : Bool;
   END_VAR
   VAR
      "CRANE STATE" : Int;
      "ENTRY N TRIG" : Bool;
      "EXIT N TRIG" : Bool;
      side : Int;
      "FREE TARGET" : Int;
      "TON-STATE-20" : TON_TIME;
      "TON-STATE-30" : TON_TIME;
      "TON-STATE-50" : TON_TIME;
      "RACK MANAGMENT_Instance" : "RACK MANAGMENT";
      warehouseFull : Bool;
      "location assigned" : Bool;
      "TON-STATE-70" : TON_TIME;
      RetrieveSide : Int;
      RetrieveLocationAssigned : Bool;
      RetrieveTarget : Int;
      "TON-STATE-100" : TON_TIME;
      "TON-STATE-120" : TON_TIME;
      "TON-STATE-140" : TON_TIME;
      "TON-STATE-160" : TON_TIME;
      "maintenance p trig" : Bool;
      "maintenance n trig" : Bool;
      "MAINTENANCE MODE" : Bool;
      "OLD STATE" : Int;
      "FAILURE DETECTION" : TON_TIME;
      "TON-STATE-130" : TON_TIME;
   END_VAR
   VAR_TEMP   // added for the SCL form of the ladder/FBD networks
      _w1 : Bool;
      _w2 : Bool;
      _w3 : Bool;
      _w4 : Bool;
   END_VAR
BEGIN

REGION Network 1
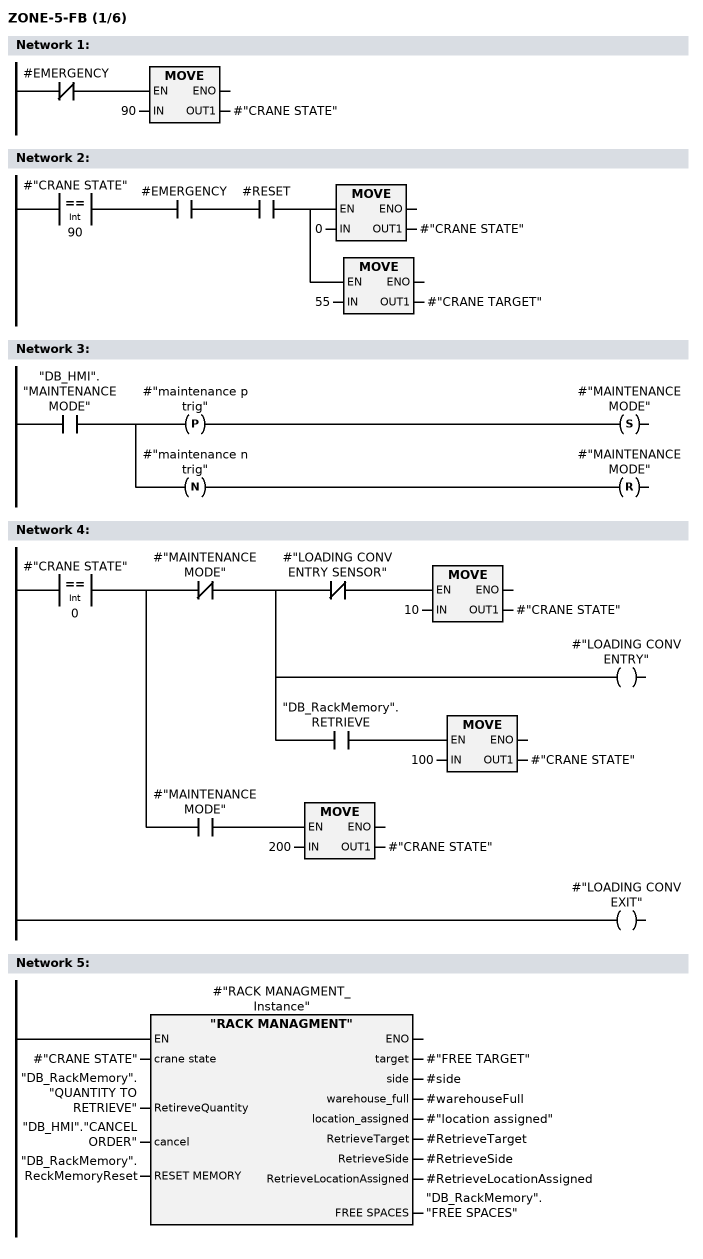
   RUNG wire#powerrail
      I_Contact( #EMERGENCY )
      Move(in := 90, out1 => #"CRANE STATE")
   END_RUNG
   // the same network as SCL:
   IF NOT #EMERGENCY THEN #"CRANE STATE" := 90; END_IF;
END_REGION

REGION Network 2
   RUNG wire#powerrail
      { S7_Templates := "SrcType := Int" } EQ_Contact(in1 := #"CRANE STATE", in2 := 90)
      Contact( #EMERGENCY )
      Contact( #RESET )
      wire#w1
      Move(in := 0, out1 => #"CRANE STATE")
   END_RUNG
   RUNG wire#w1
      Move(in := 55, out1 => #"CRANE TARGET")
   END_RUNG
   // the same network as SCL:
   #_w1 := (#"CRANE STATE" = 90) AND #EMERGENCY AND #RESET;
   IF #_w1 THEN
       #"CRANE STATE" := 0;
       #"CRANE TARGET" := 55;
   END_IF;
END_REGION

REGION Network 3
   RUNG wire#powerrail
      Contact( "DB_HMI"."MAINTENANCE MODE" )
      wire#w1
      P_Trig( #"maintenance p trig" )
      S_Coil( #"MAINTENANCE MODE" )
   END_RUNG
   RUNG wire#w1
      N_Trig( #"maintenance n trig" )
      R_Coil( #"MAINTENANCE MODE" )
   END_RUNG
   // the same network as SCL:
   #_w1 := "DB_HMI"."MAINTENANCE MODE" AND NOT #"maintenance p trig";   // rising edge
   #"maintenance p trig" := "DB_HMI"."MAINTENANCE MODE";
   IF #_w1 THEN #"MAINTENANCE MODE" := TRUE; END_IF;
   #_w2 := NOT "DB_HMI"."MAINTENANCE MODE" AND #"maintenance n trig";   // falling edge
   #"maintenance n trig" := "DB_HMI"."MAINTENANCE MODE";
   IF #_w2 THEN #"MAINTENANCE MODE" := FALSE; END_IF;
END_REGION

REGION Network 4
   RUNG wire#powerrail
      { S7_Templates := "SrcType := Int" } EQ_Contact(in1 := #"CRANE STATE", in2 := 0)
      wire#w1
      I_Contact( #"MAINTENANCE MODE" )
      wire#w2
      I_Contact( #"LOADING CONV ENTRY SENSOR" )
      Move(in := 10, out1 => #"CRANE STATE")
   END_RUNG
   RUNG wire#w2
      Coil( #"LOADING CONV ENTRY" )
   END_RUNG
   RUNG wire#w2
      Contact( "DB_RackMemory".RETRIEVE )
      Move(in := 100, out1 => #"CRANE STATE")
   END_RUNG
   RUNG wire#w1
      Contact( #"MAINTENANCE MODE" )
      Move(in := 200, out1 => #"CRANE STATE")
   END_RUNG
   RUNG wire#powerrail
      Coil( #"LOADING CONV EXIT" )
   END_RUNG
   // the same network as SCL:
   #_w1 := #"CRANE STATE" = 0;
   #_w2 := #_w1 AND NOT #"MAINTENANCE MODE";
   IF #_w2 AND NOT #"LOADING CONV ENTRY SENSOR" THEN #"CRANE STATE" := 10; END_IF;
   #"LOADING CONV ENTRY" := #_w2;
   IF #_w2 AND "DB_RackMemory".RETRIEVE THEN #"CRANE STATE" := 100; END_IF;
   IF #_w1 AND #"MAINTENANCE MODE" THEN #"CRANE STATE" := 200; END_IF;
   #"LOADING CONV EXIT" := TRUE;
END_REGION

REGION Network 5
   RUNG wire#powerrail
      #"RACK MANAGMENT_Instance"("crane state" := #"CRANE STATE", RetireveQuantity := "DB_RackMemory"."QUANTITY TO RETRIEVE", cancel := "DB_HMI"."CANCEL ORDER", "RESET MEMORY" := "DB_RackMemory".ReckMemoryReset, target => #"FREE TARGET", side => #side, warehouse_full => #warehouseFull, location_assigned => #"location assigned", RetrieveTarget => #RetrieveTarget, RetrieveSide => #RetrieveSide, RetrieveLocationAssigned => #RetrieveLocationAssigned, "FREE SPACES" => "DB_RackMemory"."FREE SPACES")
   END_RUNG
   // the same network as SCL:
   #"RACK MANAGMENT_Instance"("crane state" := #"CRANE STATE",   // "RACK MANAGMENT"
                           RetireveQuantity := "DB_RackMemory"."QUANTITY TO RETRIEVE",
                           cancel := "DB_HMI"."CANCEL ORDER",
                           "RESET MEMORY" := "DB_RackMemory".ReckMemoryReset,
                           target => #"FREE TARGET",
                           side => #side,
                           warehouse_full => #warehouseFull,
                           location_assigned => #"location assigned",
                           RetrieveTarget => #RetrieveTarget,
                           RetrieveSide => #RetrieveSide,
                           RetrieveLocationAssigned => #RetrieveLocationAssigned,
                           "FREE SPACES" => "DB_RackMemory"."FREE SPACES");
END_REGION

REGION Network 6